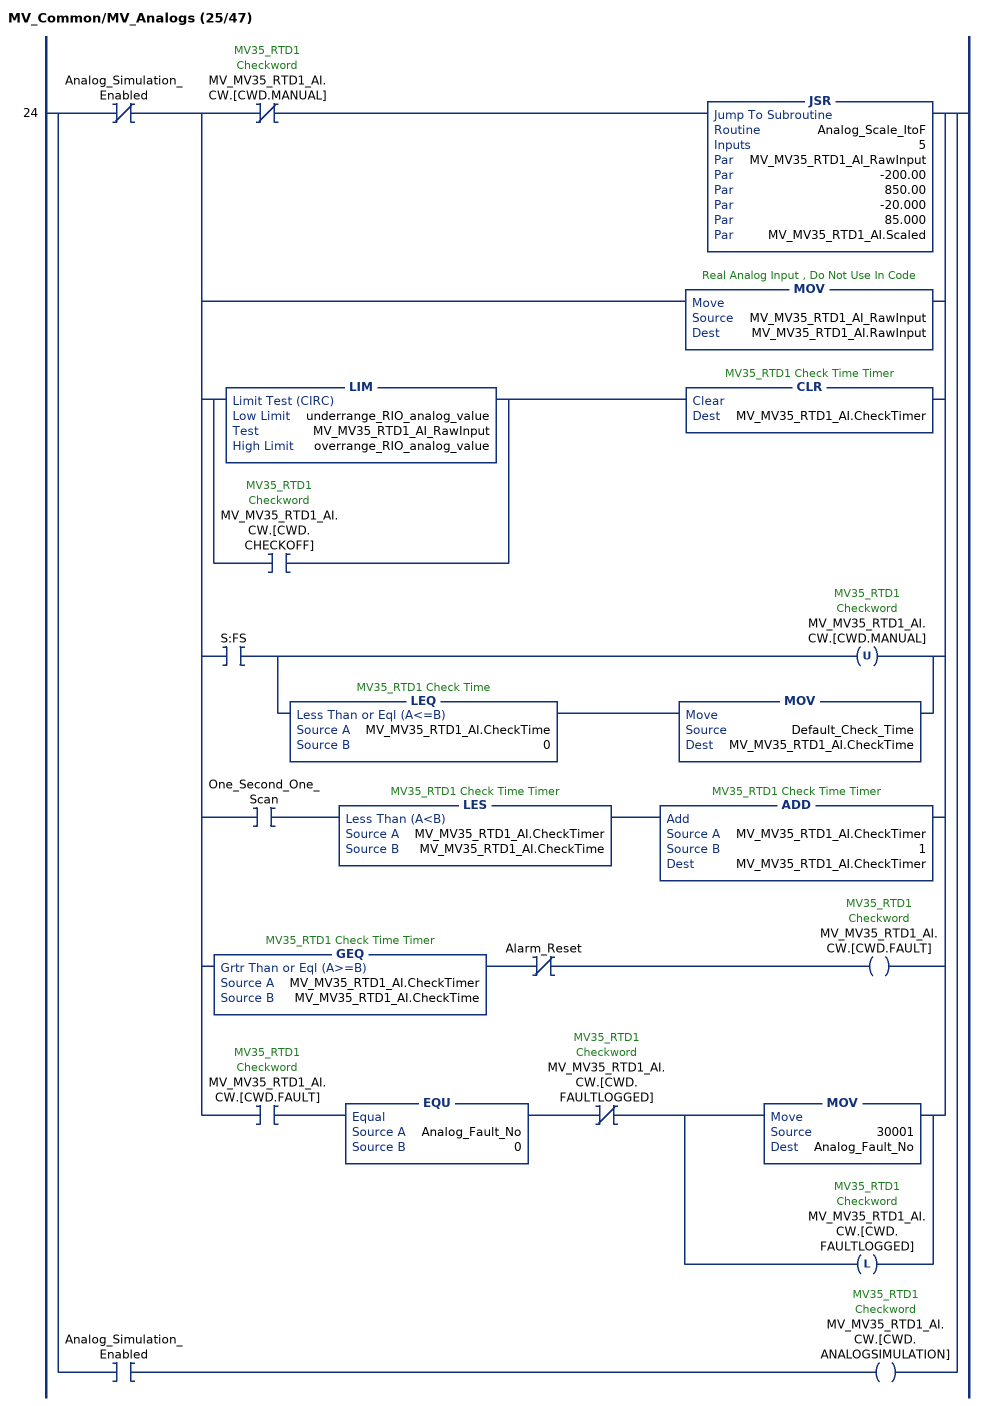
   24: [XIO(Analog_Simulation_Enabled) [XIO(MV_MV35_RTD1_AI.CW.[CWD.MANUAL]) JSR(Analog_Scale_ItoF,5,MV_MV35_RTD1_AI_RawInput,-200.00,850.00,-20.000,85.000,MV_MV35_RTD1_AI.Scaled) ,MOV(MV_MV35_RTD1_AI_RawInput,MV_MV35_RTD1_AI.RawInput) ,[LIM(underrange_RIO_analog_value,MV_MV35_RTD1_AI_RawInput,overrange_RIO_analog_value) ,XIC(MV_MV35_RTD1_AI.CW.[CWD.CHECKOFF]) ] CLR(MV_MV35_RTD1_AI.CheckTimer) ,XIC(S:FS) [OTU(MV_MV35_RTD1_AI.CW.[CWD.MANUAL]) ,LEQ(MV_MV35_RTD1_AI.CheckTime,0) MOV(Default_Check_Time,MV_MV35_RTD1_AI.CheckTime) ] ,XIC(One_Second_One_Scan) LES(MV_MV35_RTD1_AI.CheckTimer,MV_MV35_RTD1_AI.CheckTime) ADD(MV_MV35_RTD1_AI.CheckTimer,1,MV_MV35_RTD1_AI.CheckTimer) ,GEQ(MV_MV35_RTD1_AI.CheckTimer,MV_MV35_RTD1_AI.CheckTime) XIO(Alarm_Reset) OTE(MV_MV35_RTD1_AI.CW.[CWD.FAULT]) ,XIC(MV_MV35_RTD1_AI.CW.[CWD.FAULT]) EQU(Analog_Fault_No,0) XIO(MV_MV35_RTD1_AI.CW.[CWD.FAULTLOGGED]) [MOV(30001,Analog_Fault_No) ,OTL(MV_MV35_RTD1_AI.CW.[CWD.FAULTLOGGED]) ] ] ,XIC(Analog_Simulation_Enabled) OTE(MV_MV35_RTD1_AI.CW.[CWD.ANALOGSIMULATION]) ];
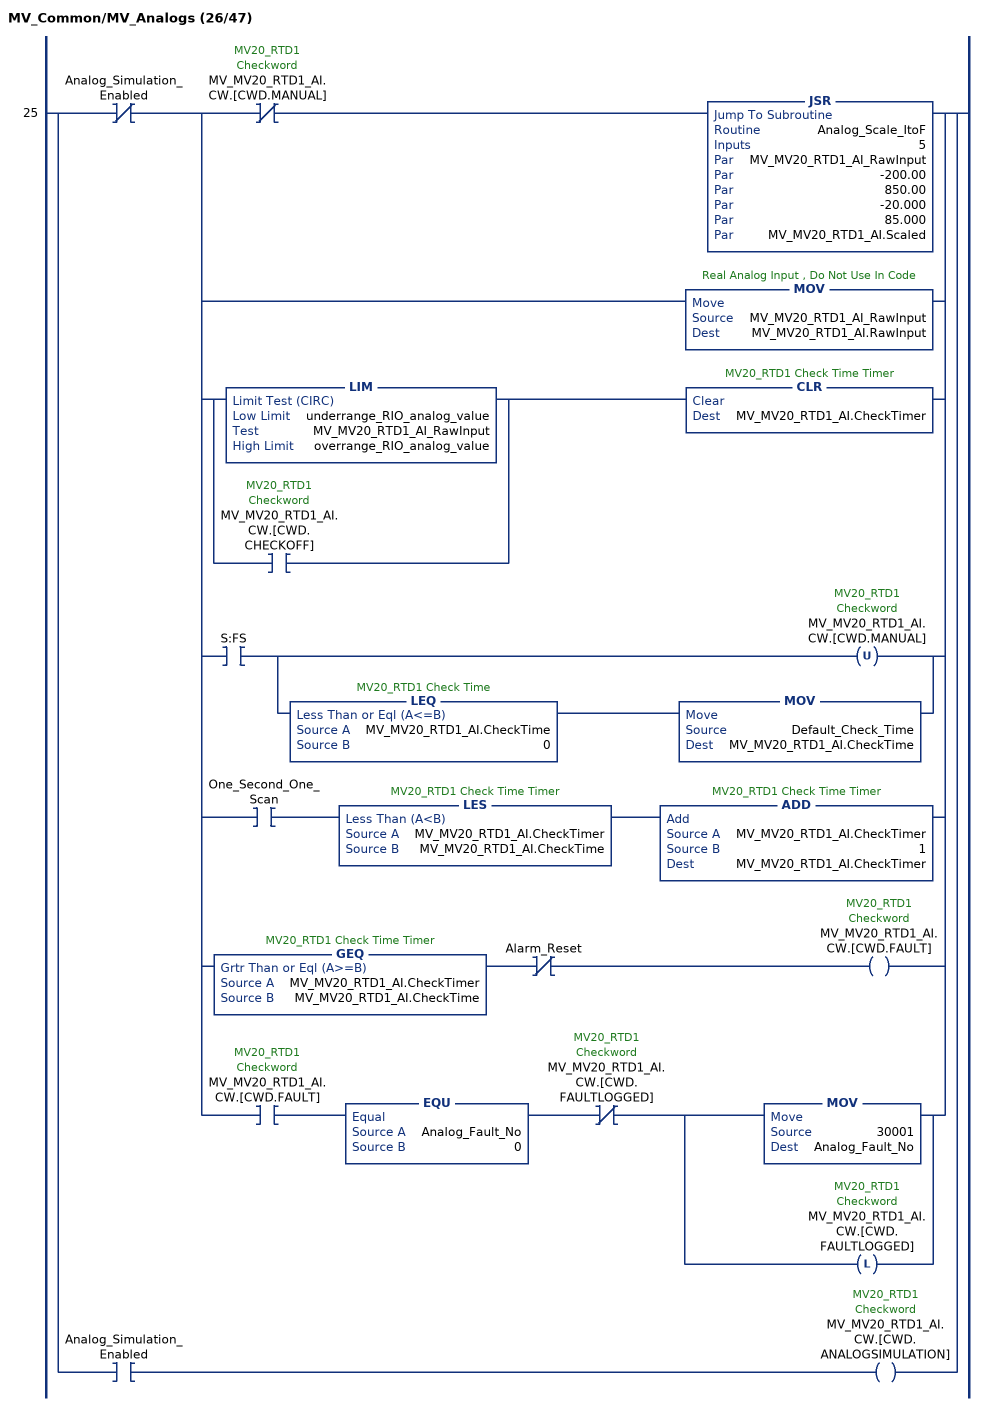
   25: [XIO(Analog_Simulation_Enabled) [XIO(MV_MV20_RTD1_AI.CW.[CWD.MANUAL]) JSR(Analog_Scale_ItoF,5,MV_MV20_RTD1_AI_RawInput,-200.00,850.00,-20.000,85.000,MV_MV20_RTD1_AI.Scaled) ,MOV(MV_MV20_RTD1_AI_RawInput,MV_MV20_RTD1_AI.RawInput) ,[LIM(underrange_RIO_analog_value,MV_MV20_RTD1_AI_RawInput,overrange_RIO_analog_value) ,XIC(MV_MV20_RTD1_AI.CW.[CWD.CHECKOFF]) ] CLR(MV_MV20_RTD1_AI.CheckTimer) ,XIC(S:FS) [OTU(MV_MV20_RTD1_AI.CW.[CWD.MANUAL]) ,LEQ(MV_MV20_RTD1_AI.CheckTime,0) MOV(Default_Check_Time,MV_MV20_RTD1_AI.CheckTime) ] ,XIC(One_Second_One_Scan) LES(MV_MV20_RTD1_AI.CheckTimer,MV_MV20_RTD1_AI.CheckTime) ADD(MV_MV20_RTD1_AI.CheckTimer,1,MV_MV20_RTD1_AI.CheckTimer) ,GEQ(MV_MV20_RTD1_AI.CheckTimer,MV_MV20_RTD1_AI.CheckTime) XIO(Alarm_Reset) OTE(MV_MV20_RTD1_AI.CW.[CWD.FAULT]) ,XIC(MV_MV20_RTD1_AI.CW.[CWD.FAULT]) EQU(Analog_Fault_No,0) XIO(MV_MV20_RTD1_AI.CW.[CWD.FAULTLOGGED]) [MOV(30001,Analog_Fault_No) ,OTL(MV_MV20_RTD1_AI.CW.[CWD.FAULTLOGGED]) ] ] ,XIC(Analog_Simulation_Enabled) OTE(MV_MV20_RTD1_AI.CW.[CWD.ANALOGSIMULATION]) ];
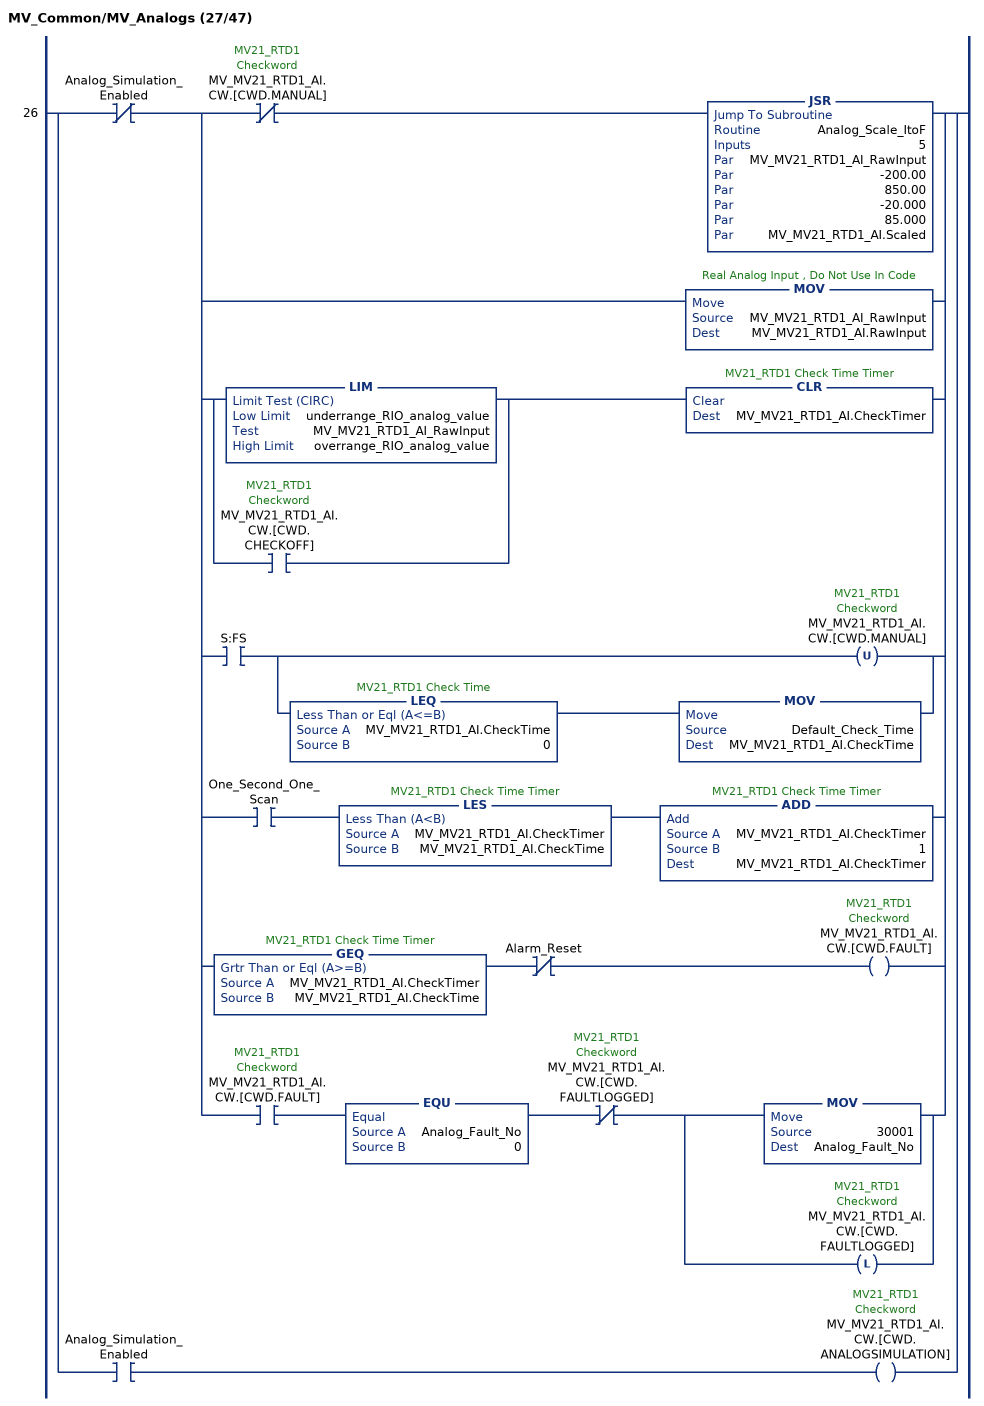
   26: [XIO(Analog_Simulation_Enabled) [XIO(MV_MV21_RTD1_AI.CW.[CWD.MANUAL]) JSR(Analog_Scale_ItoF,5,MV_MV21_RTD1_AI_RawInput,-200.00,850.00,-20.000,85.000,MV_MV21_RTD1_AI.Scaled) ,MOV(MV_MV21_RTD1_AI_RawInput,MV_MV21_RTD1_AI.RawInput) ,[LIM(underrange_RIO_analog_value,MV_MV21_RTD1_AI_RawInput,overrange_RIO_analog_value) ,XIC(MV_MV21_RTD1_AI.CW.[CWD.CHECKOFF]) ] CLR(MV_MV21_RTD1_AI.CheckTimer) ,XIC(S:FS) [OTU(MV_MV21_RTD1_AI.CW.[CWD.MANUAL]) ,LEQ(MV_MV21_RTD1_AI.CheckTime,0) MOV(Default_Check_Time,MV_MV21_RTD1_AI.CheckTime) ] ,XIC(One_Second_One_Scan) LES(MV_MV21_RTD1_AI.CheckTimer,MV_MV21_RTD1_AI.CheckTime) ADD(MV_MV21_RTD1_AI.CheckTimer,1,MV_MV21_RTD1_AI.CheckTimer) ,GEQ(MV_MV21_RTD1_AI.CheckTimer,MV_MV21_RTD1_AI.CheckTime) XIO(Alarm_Reset) OTE(MV_MV21_RTD1_AI.CW.[CWD.FAULT]) ,XIC(MV_MV21_RTD1_AI.CW.[CWD.FAULT]) EQU(Analog_Fault_No,0) XIO(MV_MV21_RTD1_AI.CW.[CWD.FAULTLOGGED]) [MOV(30001,Analog_Fault_No) ,OTL(MV_MV21_RTD1_AI.CW.[CWD.FAULTLOGGED]) ] ] ,XIC(Analog_Simulation_Enabled) OTE(MV_MV21_RTD1_AI.CW.[CWD.ANALOGSIMULATION]) ];
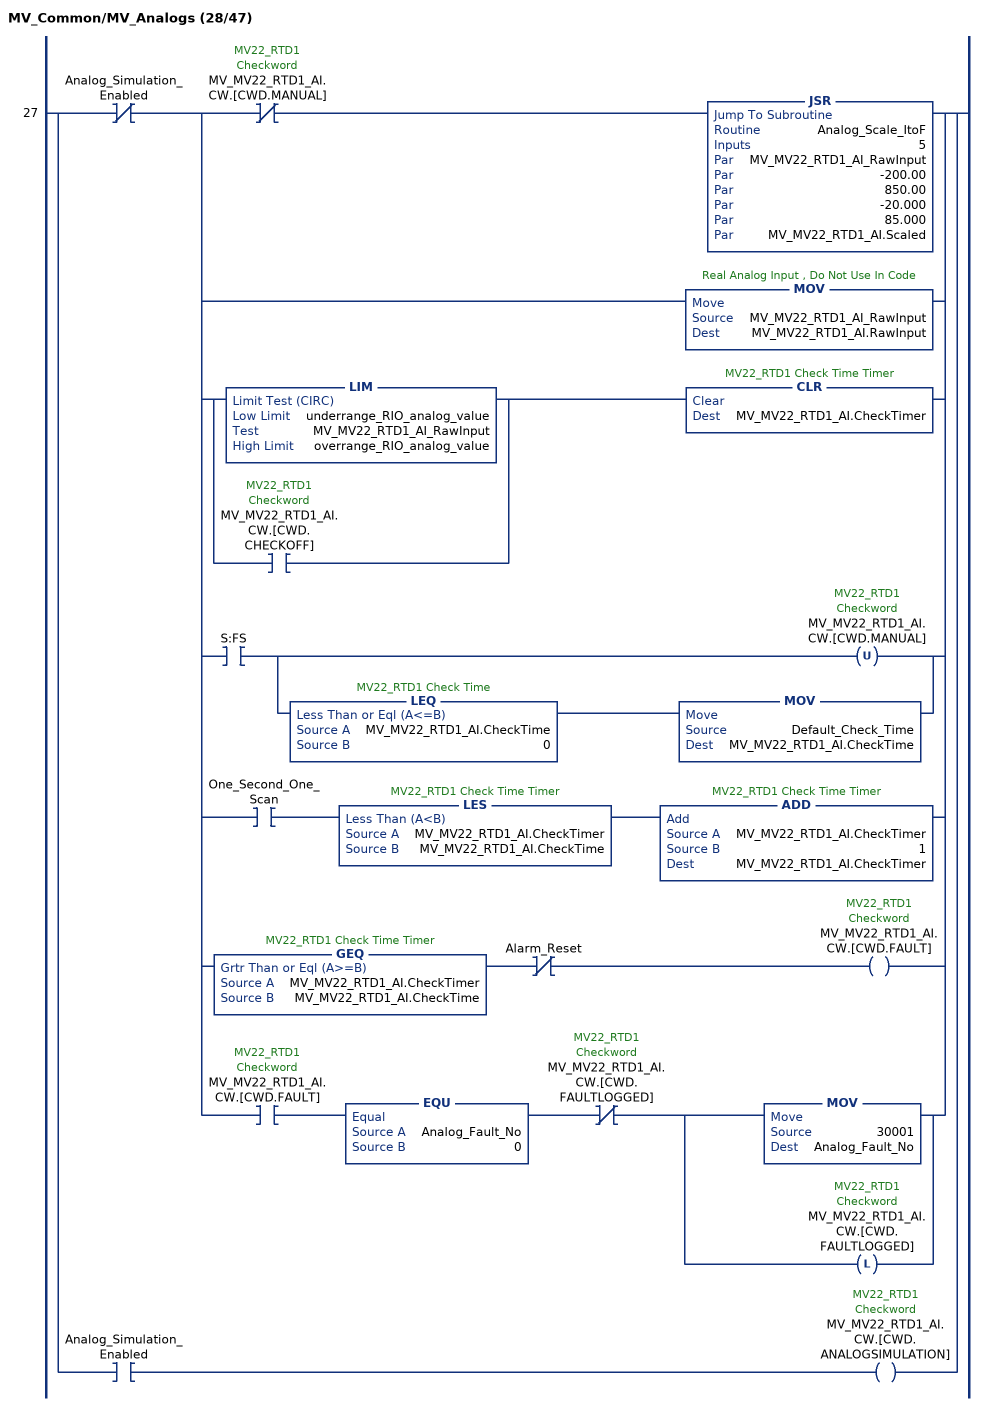
   27: [XIO(Analog_Simulation_Enabled) [XIO(MV_MV22_RTD1_AI.CW.[CWD.MANUAL]) JSR(Analog_Scale_ItoF,5,MV_MV22_RTD1_AI_RawInput,-200.00,850.00,-20.000,85.000,MV_MV22_RTD1_AI.Scaled) ,MOV(MV_MV22_RTD1_AI_RawInput,MV_MV22_RTD1_AI.RawInput) ,[LIM(underrange_RIO_analog_value,MV_MV22_RTD1_AI_RawInput,overrange_RIO_analog_value) ,XIC(MV_MV22_RTD1_AI.CW.[CWD.CHECKOFF]) ] CLR(MV_MV22_RTD1_AI.CheckTimer) ,XIC(S:FS) [OTU(MV_MV22_RTD1_AI.CW.[CWD.MANUAL]) ,LEQ(MV_MV22_RTD1_AI.CheckTime,0) MOV(Default_Check_Time,MV_MV22_RTD1_AI.CheckTime) ] ,XIC(One_Second_One_Scan) LES(MV_MV22_RTD1_AI.CheckTimer,MV_MV22_RTD1_AI.CheckTime) ADD(MV_MV22_RTD1_AI.CheckTimer,1,MV_MV22_RTD1_AI.CheckTimer) ,GEQ(MV_MV22_RTD1_AI.CheckTimer,MV_MV22_RTD1_AI.CheckTime) XIO(Alarm_Reset) OTE(MV_MV22_RTD1_AI.CW.[CWD.FAULT]) ,XIC(MV_MV22_RTD1_AI.CW.[CWD.FAULT]) EQU(Analog_Fault_No,0) XIO(MV_MV22_RTD1_AI.CW.[CWD.FAULTLOGGED]) [MOV(30001,Analog_Fault_No) ,OTL(MV_MV22_RTD1_AI.CW.[CWD.FAULTLOGGED]) ] ] ,XIC(Analog_Simulation_Enabled) OTE(MV_MV22_RTD1_AI.CW.[CWD.ANALOGSIMULATION]) ];
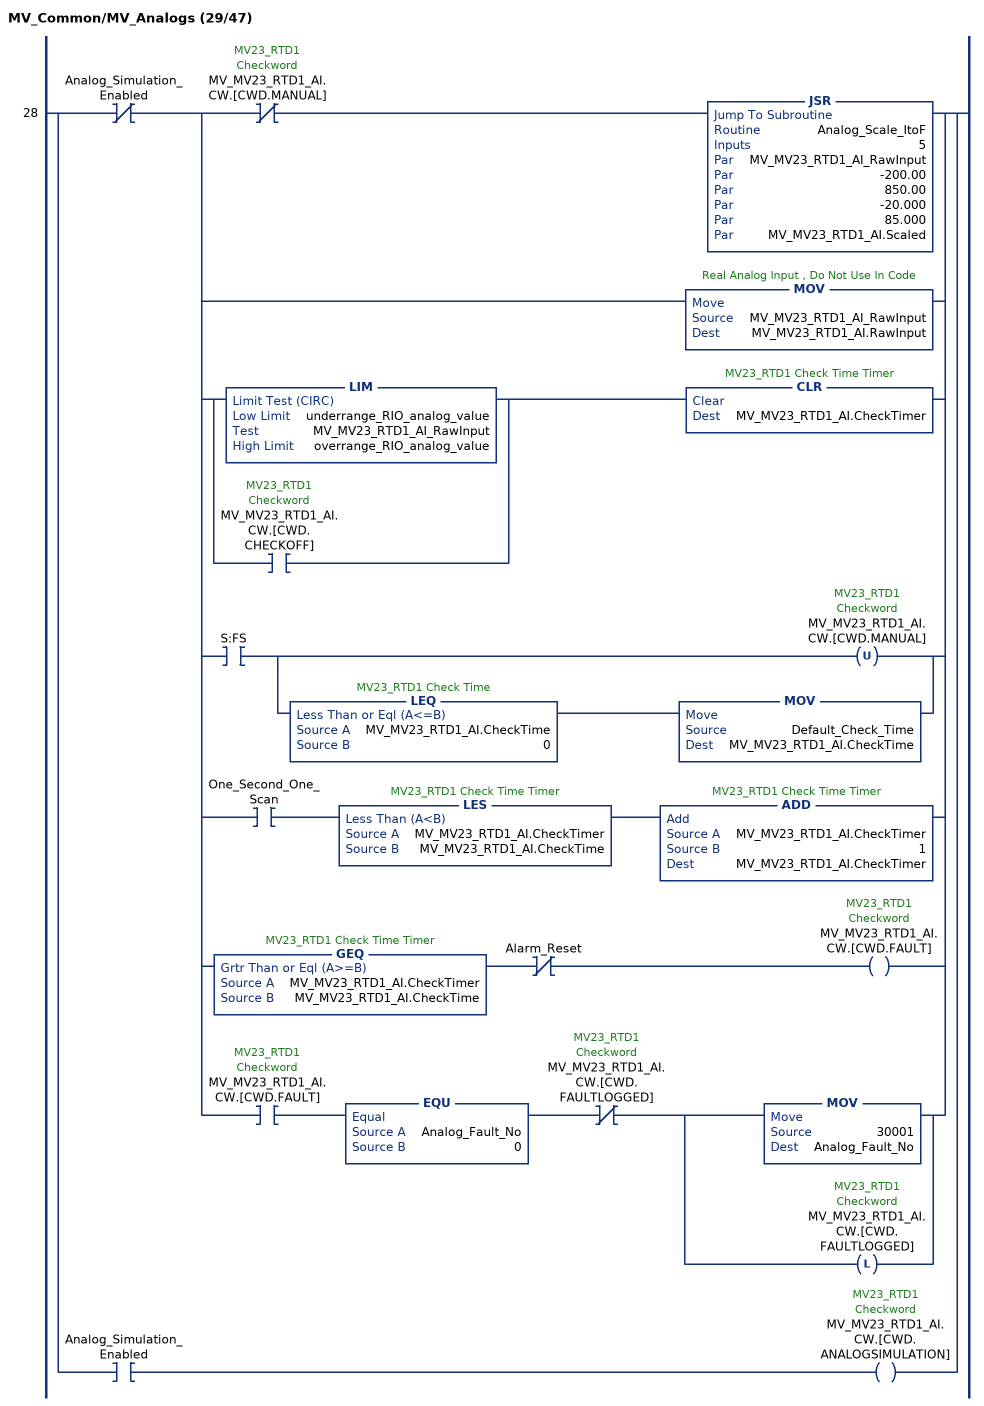
   28: [XIO(Analog_Simulation_Enabled) [XIO(MV_MV23_RTD1_AI.CW.[CWD.MANUAL]) JSR(Analog_Scale_ItoF,5,MV_MV23_RTD1_AI_RawInput,-200.00,850.00,-20.000,85.000,MV_MV23_RTD1_AI.Scaled) ,MOV(MV_MV23_RTD1_AI_RawInput,MV_MV23_RTD1_AI.RawInput) ,[LIM(underrange_RIO_analog_value,MV_MV23_RTD1_AI_RawInput,overrange_RIO_analog_value) ,XIC(MV_MV23_RTD1_AI.CW.[CWD.CHECKOFF]) ] CLR(MV_MV23_RTD1_AI.CheckTimer) ,XIC(S:FS) [OTU(MV_MV23_RTD1_AI.CW.[CWD.MANUAL]) ,LEQ(MV_MV23_RTD1_AI.CheckTime,0) MOV(Default_Check_Time,MV_MV23_RTD1_AI.CheckTime) ] ,XIC(One_Second_One_Scan) LES(MV_MV23_RTD1_AI.CheckTimer,MV_MV23_RTD1_AI.CheckTime) ADD(MV_MV23_RTD1_AI.CheckTimer,1,MV_MV23_RTD1_AI.CheckTimer) ,GEQ(MV_MV23_RTD1_AI.CheckTimer,MV_MV23_RTD1_AI.CheckTime) XIO(Alarm_Reset) OTE(MV_MV23_RTD1_AI.CW.[CWD.FAULT]) ,XIC(MV_MV23_RTD1_AI.CW.[CWD.FAULT]) EQU(Analog_Fault_No,0) XIO(MV_MV23_RTD1_AI.CW.[CWD.FAULTLOGGED]) [MOV(30001,Analog_Fault_No) ,OTL(MV_MV23_RTD1_AI.CW.[CWD.FAULTLOGGED]) ] ] ,XIC(Analog_Simulation_Enabled) OTE(MV_MV23_RTD1_AI.CW.[CWD.ANALOGSIMULATION]) ];
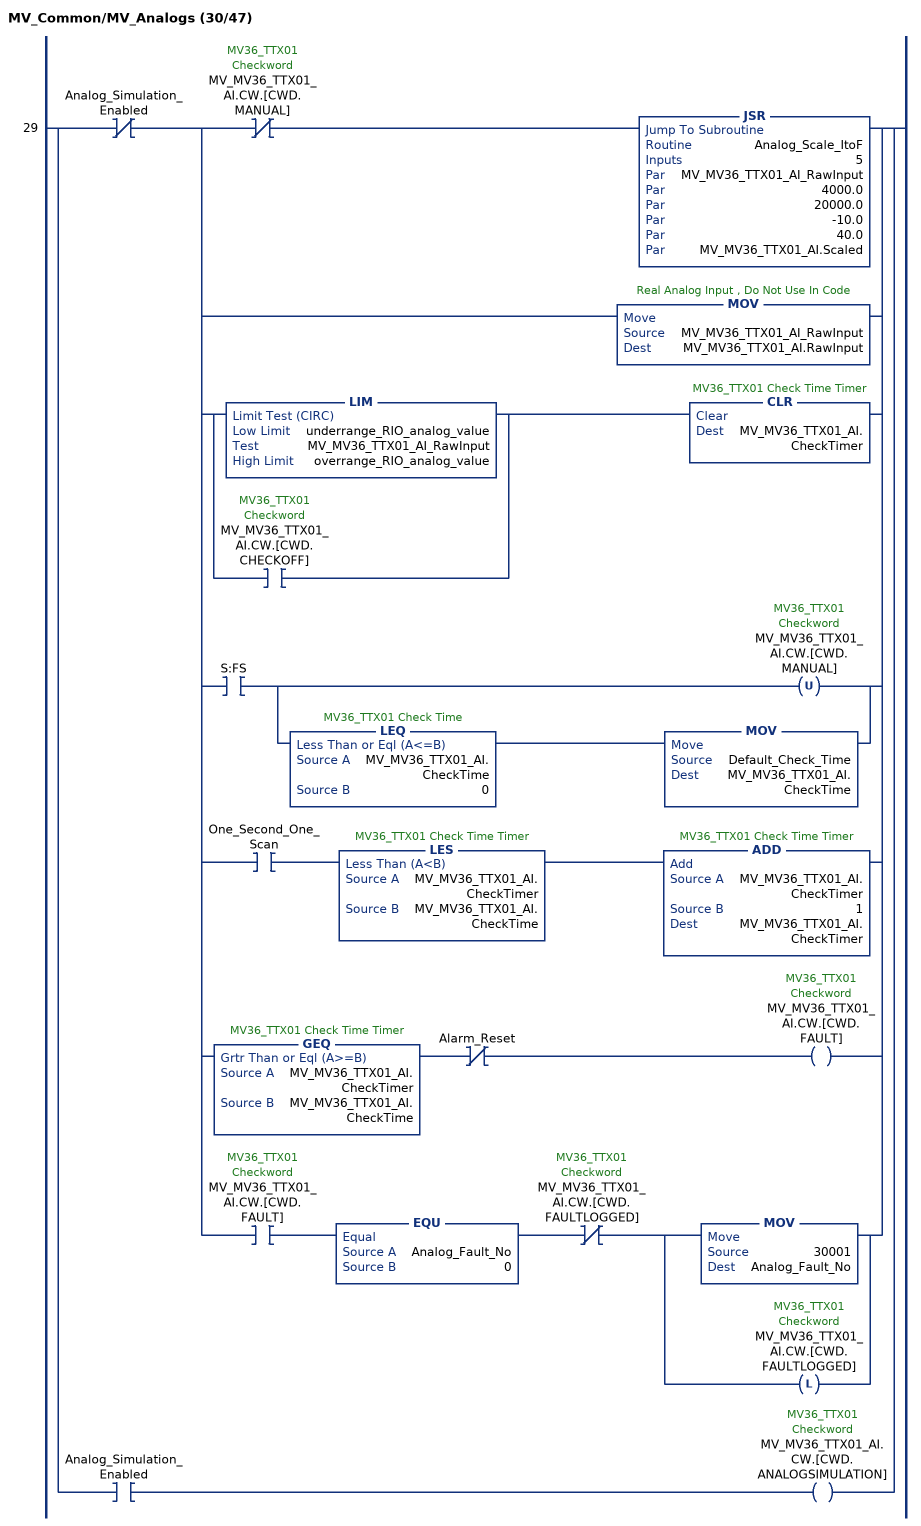
   29: [XIO(Analog_Simulation_Enabled) [XIO(MV_MV36_TTX01_AI.CW.[CWD.MANUAL]) JSR(Analog_Scale_ItoF,5,MV_MV36_TTX01_AI_RawInput,4000.0,20000.0,-10.0,40.0,MV_MV36_TTX01_AI.Scaled) ,MOV(MV_MV36_TTX01_AI_RawInput,MV_MV36_TTX01_AI.RawInput) ,[LIM(underrange_RIO_analog_value,MV_MV36_TTX01_AI_RawInput,overrange_RIO_analog_value) ,XIC(MV_MV36_TTX01_AI.CW.[CWD.CHECKOFF]) ] CLR(MV_MV36_TTX01_AI.CheckTimer) ,XIC(S:FS) [OTU(MV_MV36_TTX01_AI.CW.[CWD.MANUAL]) ,LEQ(MV_MV36_TTX01_AI.CheckTime,0) MOV(Default_Check_Time,MV_MV36_TTX01_AI.CheckTime) ] ,XIC(One_Second_One_Scan) LES(MV_MV36_TTX01_AI.CheckTimer,MV_MV36_TTX01_AI.CheckTime) ADD(MV_MV36_TTX01_AI.CheckTimer,1,MV_MV36_TTX01_AI.CheckTimer) ,GEQ(MV_MV36_TTX01_AI.CheckTimer,MV_MV36_TTX01_AI.CheckTime) XIO(Alarm_Reset) OTE(MV_MV36_TTX01_AI.CW.[CWD.FAULT]) ,XIC(MV_MV36_TTX01_AI.CW.[CWD.FAULT]) EQU(Analog_Fault_No,0) XIO(MV_MV36_TTX01_AI.CW.[CWD.FAULTLOGGED]) [MOV(30001,Analog_Fault_No) ,OTL(MV_MV36_TTX01_AI.CW.[CWD.FAULTLOGGED]) ] ] ,XIC(Analog_Simulation_Enabled) OTE(MV_MV36_TTX01_AI.CW.[CWD.ANALOGSIMULATION]) ];
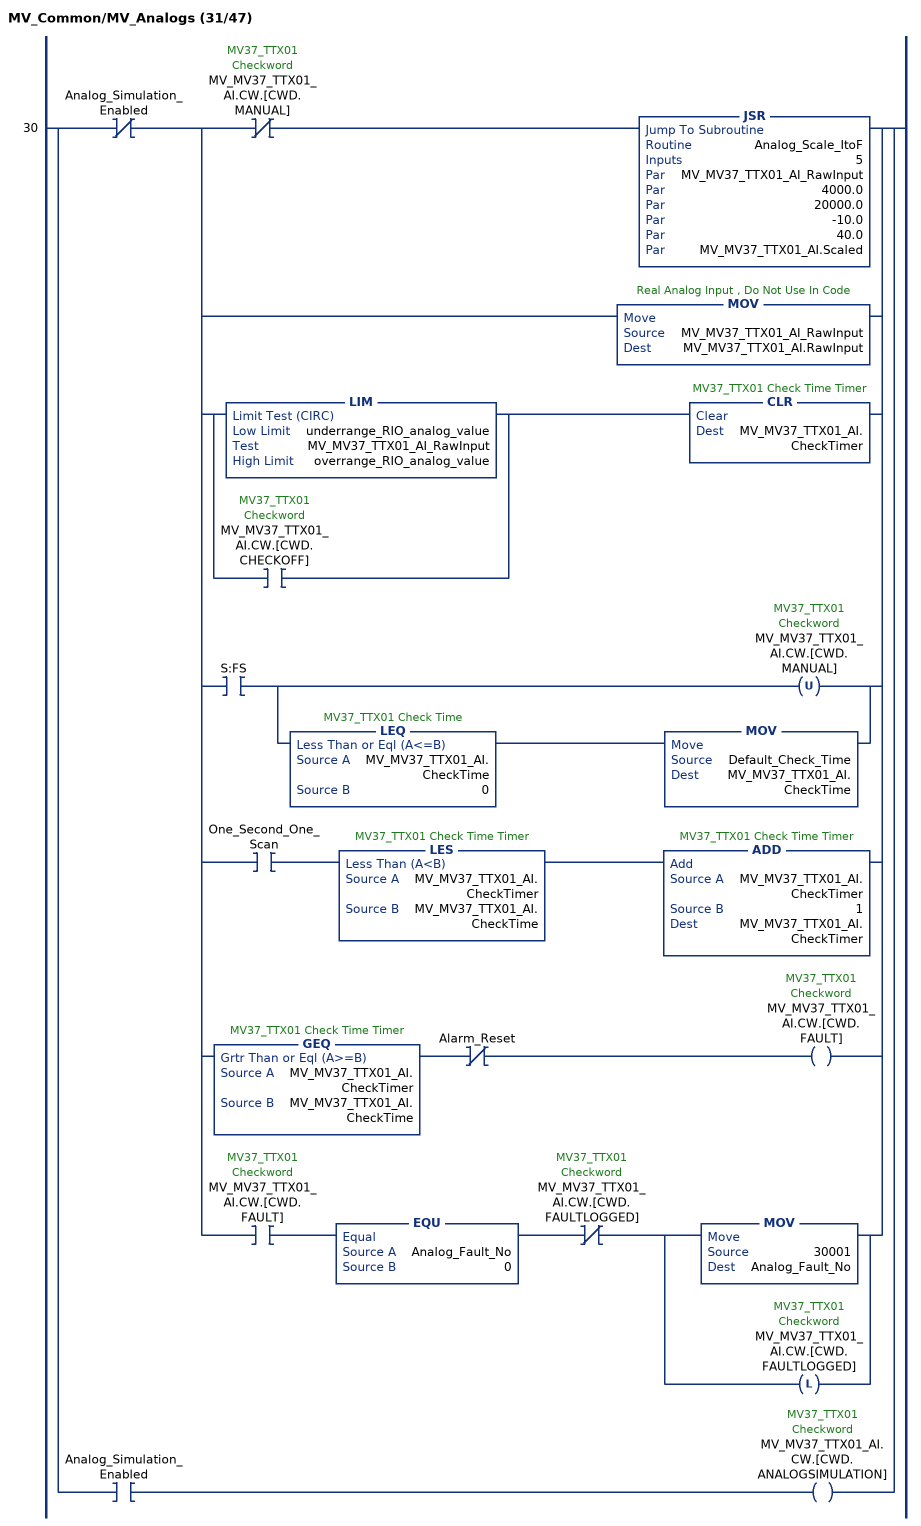
   30: [XIO(Analog_Simulation_Enabled) [XIO(MV_MV37_TTX01_AI.CW.[CWD.MANUAL]) JSR(Analog_Scale_ItoF,5,MV_MV37_TTX01_AI_RawInput,4000.0,20000.0,-10.0,40.0,MV_MV37_TTX01_AI.Scaled) ,MOV(MV_MV37_TTX01_AI_RawInput,MV_MV37_TTX01_AI.RawInput) ,[LIM(underrange_RIO_analog_value,MV_MV37_TTX01_AI_RawInput,overrange_RIO_analog_value) ,XIC(MV_MV37_TTX01_AI.CW.[CWD.CHECKOFF]) ] CLR(MV_MV37_TTX01_AI.CheckTimer) ,XIC(S:FS) [OTU(MV_MV37_TTX01_AI.CW.[CWD.MANUAL]) ,LEQ(MV_MV37_TTX01_AI.CheckTime,0) MOV(Default_Check_Time,MV_MV37_TTX01_AI.CheckTime) ] ,XIC(One_Second_One_Scan) LES(MV_MV37_TTX01_AI.CheckTimer,MV_MV37_TTX01_AI.CheckTime) ADD(MV_MV37_TTX01_AI.CheckTimer,1,MV_MV37_TTX01_AI.CheckTimer) ,GEQ(MV_MV37_TTX01_AI.CheckTimer,MV_MV37_TTX01_AI.CheckTime) XIO(Alarm_Reset) OTE(MV_MV37_TTX01_AI.CW.[CWD.FAULT]) ,XIC(MV_MV37_TTX01_AI.CW.[CWD.FAULT]) EQU(Analog_Fault_No,0) XIO(MV_MV37_TTX01_AI.CW.[CWD.FAULTLOGGED]) [MOV(30001,Analog_Fault_No) ,OTL(MV_MV37_TTX01_AI.CW.[CWD.FAULTLOGGED]) ] ] ,XIC(Analog_Simulation_Enabled) OTE(MV_MV37_TTX01_AI.CW.[CWD.ANALOGSIMULATION]) ];
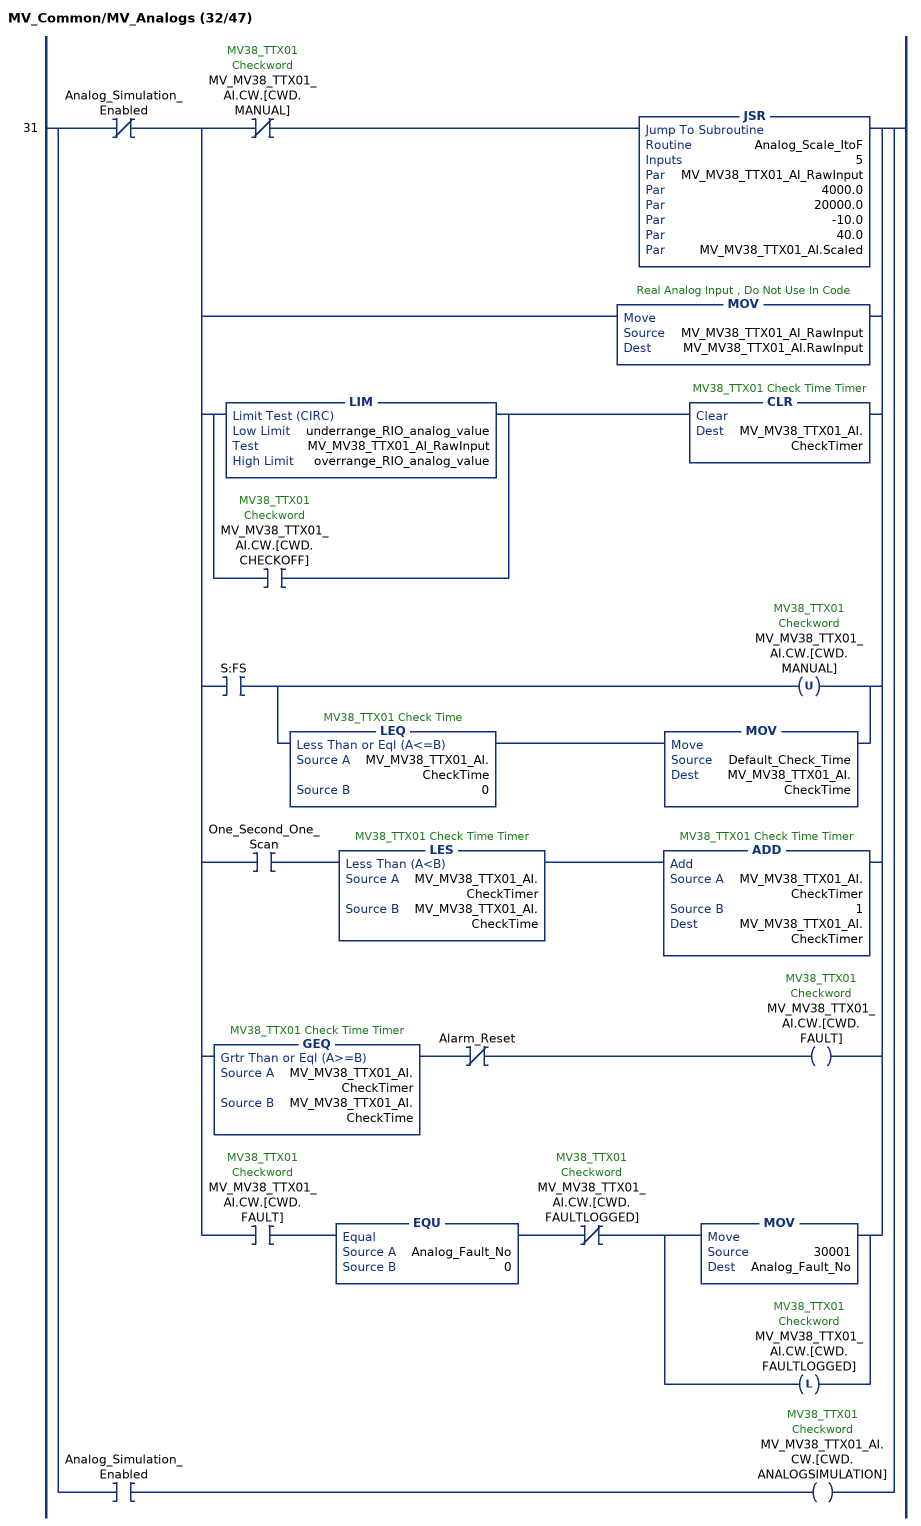
   31: [XIO(Analog_Simulation_Enabled) [XIO(MV_MV38_TTX01_AI.CW.[CWD.MANUAL]) JSR(Analog_Scale_ItoF,5,MV_MV38_TTX01_AI_RawInput,4000.0,20000.0,-10.0,40.0,MV_MV38_TTX01_AI.Scaled) ,MOV(MV_MV38_TTX01_AI_RawInput,MV_MV38_TTX01_AI.RawInput) ,[LIM(underrange_RIO_analog_value,MV_MV38_TTX01_AI_RawInput,overrange_RIO_analog_value) ,XIC(MV_MV38_TTX01_AI.CW.[CWD.CHECKOFF]) ] CLR(MV_MV38_TTX01_AI.CheckTimer) ,XIC(S:FS) [OTU(MV_MV38_TTX01_AI.CW.[CWD.MANUAL]) ,LEQ(MV_MV38_TTX01_AI.CheckTime,0) MOV(Default_Check_Time,MV_MV38_TTX01_AI.CheckTime) ] ,XIC(One_Second_One_Scan) LES(MV_MV38_TTX01_AI.CheckTimer,MV_MV38_TTX01_AI.CheckTime) ADD(MV_MV38_TTX01_AI.CheckTimer,1,MV_MV38_TTX01_AI.CheckTimer) ,GEQ(MV_MV38_TTX01_AI.CheckTimer,MV_MV38_TTX01_AI.CheckTime) XIO(Alarm_Reset) OTE(MV_MV38_TTX01_AI.CW.[CWD.FAULT]) ,XIC(MV_MV38_TTX01_AI.CW.[CWD.FAULT]) EQU(Analog_Fault_No,0) XIO(MV_MV38_TTX01_AI.CW.[CWD.FAULTLOGGED]) [MOV(30001,Analog_Fault_No) ,OTL(MV_MV38_TTX01_AI.CW.[CWD.FAULTLOGGED]) ] ] ,XIC(Analog_Simulation_Enabled) OTE(MV_MV38_TTX01_AI.CW.[CWD.ANALOGSIMULATION]) ];